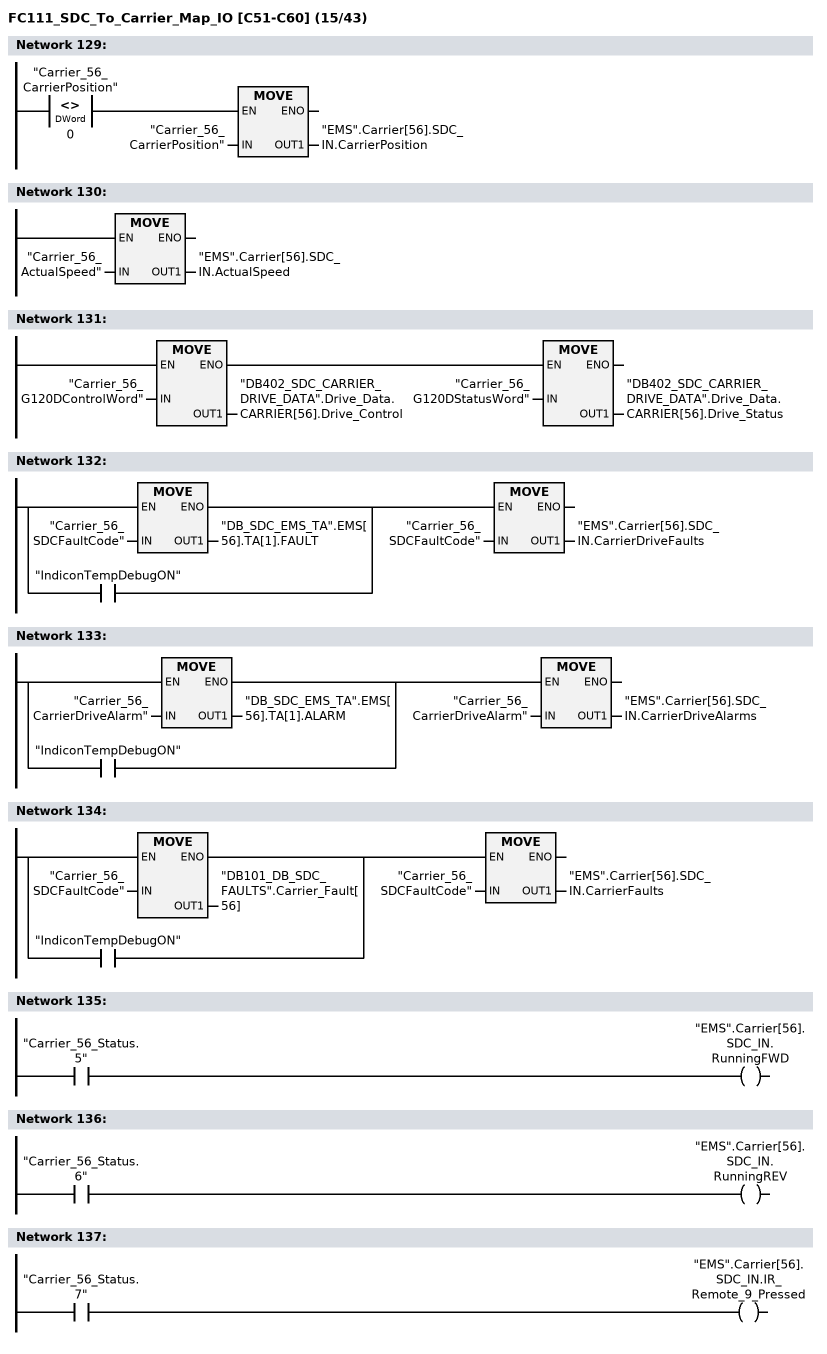
   RUNG wire#powerrail
      { S7_Templates := "SrcType := DWord" } NE_Contact(in1 := "Carrier_56_CarrierPosition", in2 := 0)
      Move(in := "Carrier_56_CarrierPosition", out1 => "EMS".Carrier[56].SDC_IN.CarrierPosition)
   END_RUNG
   // the same network as SCL:
   IF "Carrier_56_CarrierPosition" <> 0 THEN
       "EMS".Carrier[56].SDC_IN.CarrierPosition := "Carrier_56_CarrierPosition";
   END_IF;
END_REGION

REGION Network 130
   RUNG wire#powerrail
      Move(in := "Carrier_56_ActualSpeed", out1 => "EMS".Carrier[56].SDC_IN.ActualSpeed)
   END_RUNG
   // the same network as SCL:
   "EMS".Carrier[56].SDC_IN.ActualSpeed := "Carrier_56_ActualSpeed";
END_REGION

REGION Network 131
   RUNG wire#powerrail
      Move(in := "Carrier_56_G120DControlWord", out1 => "DB402_SDC_CARRIER_DRIVE_DATA".Drive_Data.CARRIER[56].Drive_Control)
      Move(in := "Carrier_56_G120DStatusWord", out1 => "DB402_SDC_CARRIER_DRIVE_DATA".Drive_Data.CARRIER[56].Drive_Status)
   END_RUNG
   // the same network as SCL:
   "DB402_SDC_CARRIER_DRIVE_DATA".Drive_Data.CARRIER[56].Drive_Control := "Carrier_56_G120DControlWord";
   "DB402_SDC_CARRIER_DRIVE_DATA".Drive_Data.CARRIER[56].Drive_Status := "Carrier_56_G120DStatusWord";
END_REGION

REGION Network 132
   RUNG wire#powerrail
      Move(in := "Carrier_56_SDCFaultCode", out1 => "DB_SDC_EMS_TA".EMS[56].TA[1].FAULT)
      wire#w1
      Move(in := "Carrier_56_SDCFaultCode", out1 => "EMS".Carrier[56].SDC_IN.CarrierDriveFaults)
   END_RUNG
   RUNG wire#powerrail
      Contact( "IndiconTempDebugON" )
   END_RUNG wire#w1
   // the same network as SCL:
   "DB_SDC_EMS_TA".EMS[56].TA[1].FAULT := "Carrier_56_SDCFaultCode";
   IF TRUE OR "IndiconTempDebugON" THEN
       "EMS".Carrier[56].SDC_IN.CarrierDriveFaults := "Carrier_56_SDCFaultCode";
   END_IF;
END_REGION

REGION Network 133
   RUNG wire#powerrail
      Move(in := "Carrier_56_CarrierDriveAlarm", out1 => "DB_SDC_EMS_TA".EMS[56].TA[1].ALARM)
      wire#w1
      Move(in := "Carrier_56_CarrierDriveAlarm", out1 => "EMS".Carrier[56].SDC_IN.CarrierDriveAlarms)
   END_RUNG
   RUNG wire#powerrail
      Contact( "IndiconTempDebugON" )
   END_RUNG wire#w1
   // the same network as SCL:
   "DB_SDC_EMS_TA".EMS[56].TA[1].ALARM := "Carrier_56_CarrierDriveAlarm";
   IF TRUE OR "IndiconTempDebugON" THEN
       "EMS".Carrier[56].SDC_IN.CarrierDriveAlarms := "Carrier_56_CarrierDriveAlarm";
   END_IF;
END_REGION

REGION Network 134
   RUNG wire#powerrail
      Move(in := "Carrier_56_SDCFaultCode", out1 => "DB101_DB_SDC_FAULTS".Carrier_Fault[56])
      wire#w1
      Move(in := "Carrier_56_SDCFaultCode", out1 => "EMS".Carrier[56].SDC_IN.CarrierFaults)
   END_RUNG
   RUNG wire#powerrail
      Contact( "IndiconTempDebugON" )
   END_RUNG wire#w1
   // the same network as SCL:
   "DB101_DB_SDC_FAULTS".Carrier_Fault[56] := "Carrier_56_SDCFaultCode";
   IF TRUE OR "IndiconTempDebugON" THEN
       "EMS".Carrier[56].SDC_IN.CarrierFaults := "Carrier_56_SDCFaultCode";
   END_IF;
END_REGION

REGION Network 135
   RUNG wire#powerrail
      Contact( "Carrier_56_Status.5" )
      Coil( "EMS".Carrier[56].SDC_IN.RunningFWD )
   END_RUNG
   // the same network as SCL:
   "EMS".Carrier[56].SDC_IN.RunningFWD := "Carrier_56_Status.5";
END_REGION

REGION Network 136
   RUNG wire#powerrail
      Contact( "Carrier_56_Status.6" )
      Coil( "EMS".Carrier[56].SDC_IN.RunningREV )
   END_RUNG
   // the same network as SCL:
   "EMS".Carrier[56].SDC_IN.RunningREV := "Carrier_56_Status.6";
END_REGION

REGION Network 137
   RUNG wire#powerrail
      Contact( "Carrier_56_Status.7" )
      Coil( "EMS".Carrier[56].SDC_IN.IR_Remote_9_Pressed )
   END_RUNG
   // the same network as SCL:
   "EMS".Carrier[56].SDC_IN.IR_Remote_9_Pressed := "Carrier_56_Status.7";
END_REGION

REGION Network 138
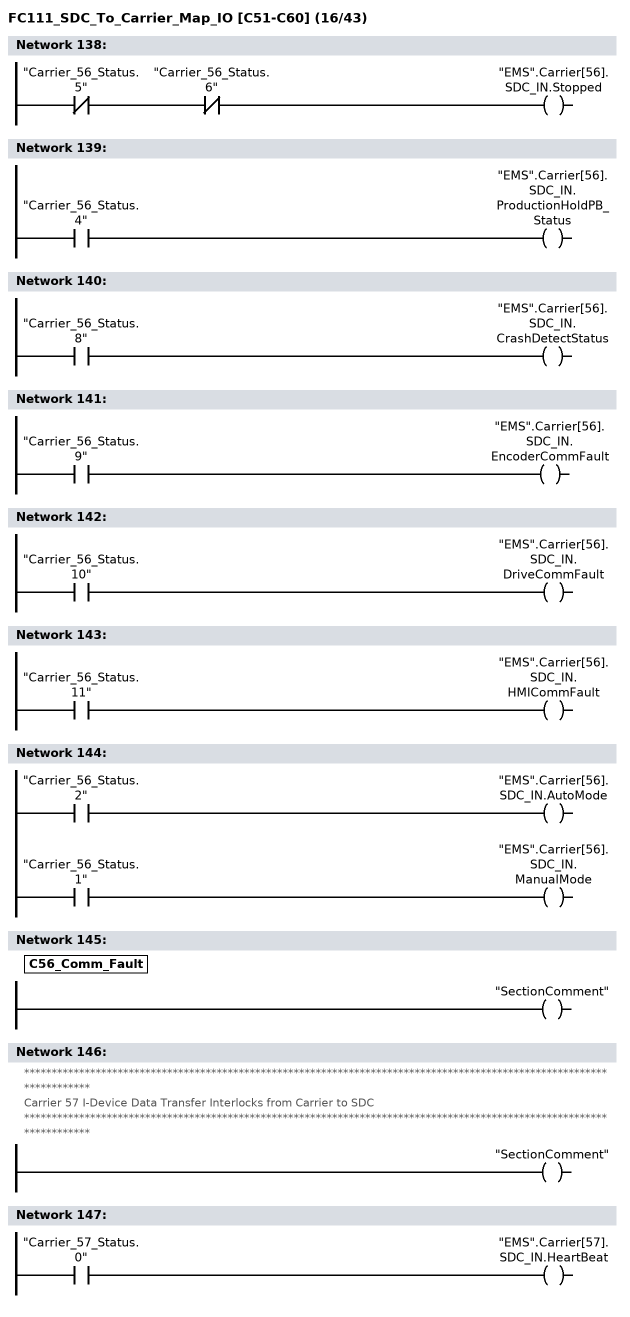
   RUNG wire#powerrail
      I_Contact( "Carrier_56_Status.5" )
      I_Contact( "Carrier_56_Status.6" )
      Coil( "EMS".Carrier[56].SDC_IN.Stopped )
   END_RUNG
   // the same network as SCL:
   "EMS".Carrier[56].SDC_IN.Stopped := NOT "Carrier_56_Status.5" AND NOT "Carrier_56_Status.6";
END_REGION

REGION Network 139
   RUNG wire#powerrail
      Contact( "Carrier_56_Status.4" )
      Coil( "EMS".Carrier[56].SDC_IN.ProductionHoldPB_Status )
   END_RUNG
   // the same network as SCL:
   "EMS".Carrier[56].SDC_IN.ProductionHoldPB_Status := "Carrier_56_Status.4";
END_REGION

REGION Network 140
   RUNG wire#powerrail
      Contact( "Carrier_56_Status.8" )
      Coil( "EMS".Carrier[56].SDC_IN.CrashDetectStatus )
   END_RUNG
   // the same network as SCL:
   "EMS".Carrier[56].SDC_IN.CrashDetectStatus := "Carrier_56_Status.8";
END_REGION

REGION Network 141
   RUNG wire#powerrail
      Contact( "Carrier_56_Status.9" )
      Coil( "EMS".Carrier[56].SDC_IN.EncoderCommFault )
   END_RUNG
   // the same network as SCL:
   "EMS".Carrier[56].SDC_IN.EncoderCommFault := "Carrier_56_Status.9";
END_REGION

REGION Network 142
   RUNG wire#powerrail
      Contact( "Carrier_56_Status.10" )
      Coil( "EMS".Carrier[56].SDC_IN.DriveCommFault )
   END_RUNG
   // the same network as SCL:
   "EMS".Carrier[56].SDC_IN.DriveCommFault := "Carrier_56_Status.10";
END_REGION

REGION Network 143
   RUNG wire#powerrail
      Contact( "Carrier_56_Status.11" )
      Coil( "EMS".Carrier[56].SDC_IN.HMICommFault )
   END_RUNG
   // the same network as SCL:
   "EMS".Carrier[56].SDC_IN.HMICommFault := "Carrier_56_Status.11";
END_REGION

REGION Network 144
   RUNG wire#powerrail
      Contact( "Carrier_56_Status.2" )
      Coil( "EMS".Carrier[56].SDC_IN.AutoMode )
   END_RUNG
   RUNG wire#powerrail
      Contact( "Carrier_56_Status.1" )
      Coil( "EMS".Carrier[56].SDC_IN.ManualMode )
   END_RUNG
   // the same network as SCL:
   "EMS".Carrier[56].SDC_IN.AutoMode := "Carrier_56_Status.2";
   "EMS".Carrier[56].SDC_IN.ManualMode := "Carrier_56_Status.1";
END_REGION

REGION Network 145
   Label( C56_Comm_Fault )
   RUNG wire#powerrail
      Coil( "SectionComment" )
   END_RUNG
   // the same network as SCL:
   C56_Comm_Fault:
   "SectionComment" := TRUE;
END_REGION

REGION Network 146
   // **********************************************************************************************************************
   // 
   // Carrier 57 I-Device Data Transfer Interlocks from Carrier to SDC
   // 
   // **********************************************************************************************************************
   RUNG wire#powerrail
      Coil( "SectionComment" )
   END_RUNG
   // the same network as SCL:
   "SectionComment" := TRUE;
END_REGION

REGION Network 147
   RUNG wire#powerrail
      Contact( "Carrier_57_Status.0" )
      Coil( "EMS".Carrier[57].SDC_IN.HeartBeat )
   END_RUNG
   // the same network as SCL:
   "EMS".Carrier[57].SDC_IN.HeartBeat := "Carrier_57_Status.0";
END_REGION

REGION Network 148
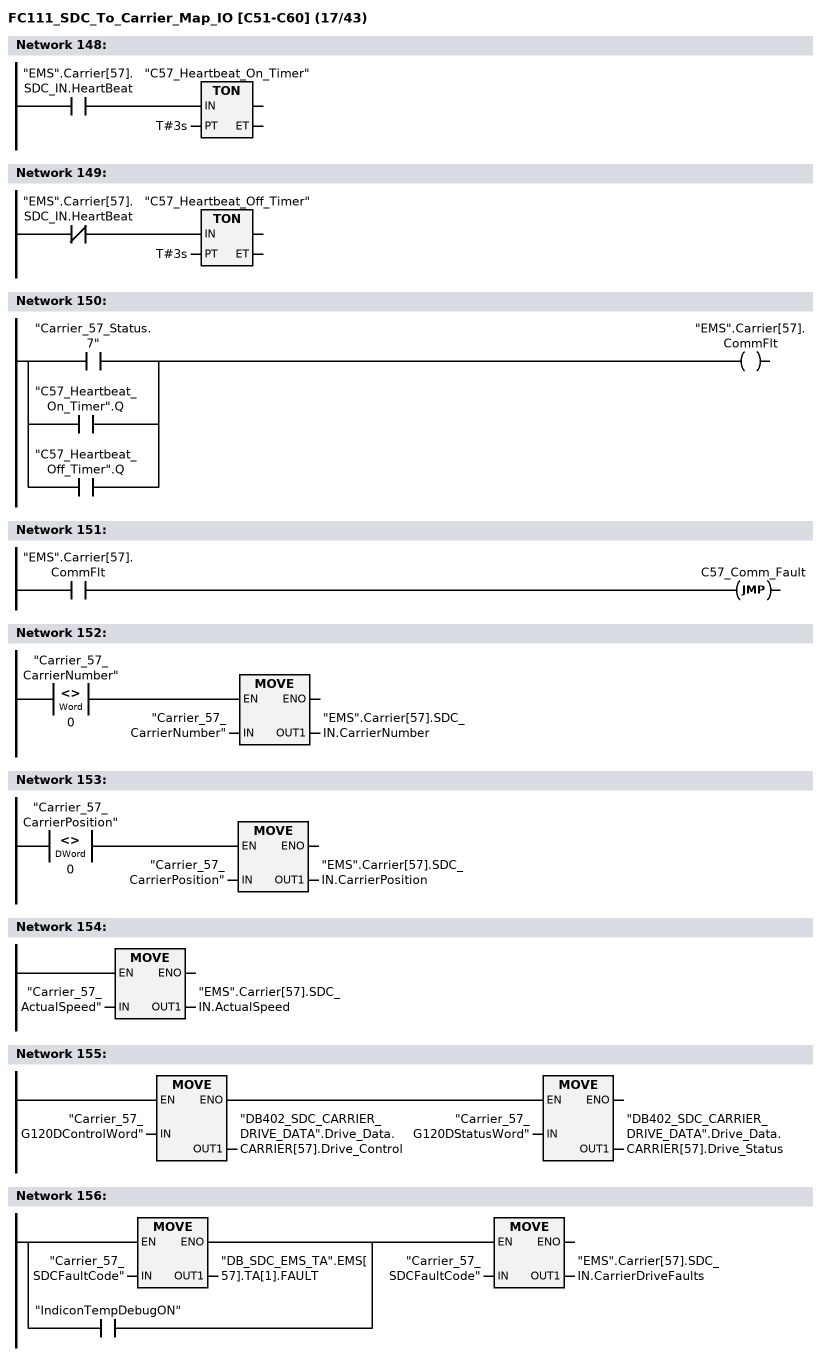
   "C57_Heartbeat_On_Timer".TON(IN := "EMS".Carrier[57].SDC_IN.HeartBeat, PT := T#3s);
END_REGION

REGION Network 149
   "C57_Heartbeat_Off_Timer".TON(IN := NOT "EMS".Carrier[57].SDC_IN.HeartBeat, PT := T#3s);
END_REGION

REGION Network 150
   RUNG wire#powerrail
      Contact( "Carrier_57_Status.7" )
      wire#w1
      Coil( "EMS".Carrier[57].CommFlt )
   END_RUNG
   RUNG wire#powerrail
      Contact( "C57_Heartbeat_On_Timer".Q )
   END_RUNG wire#w1
   RUNG wire#powerrail
      Contact( "C57_Heartbeat_Off_Timer".Q )
   END_RUNG wire#w1
   // the same network as SCL:
   "EMS".Carrier[57].CommFlt := "Carrier_57_Status.7" OR "C57_Heartbeat_On_Timer".Q OR "C57_Heartbeat_Off_Timer".Q;
END_REGION

REGION Network 151
   RUNG wire#powerrail
      Contact( "EMS".Carrier[57].CommFlt )
      JumpCoil( C57_Comm_Fault )
   END_RUNG
   // the same network as SCL:
   IF "EMS".Carrier[57].CommFlt THEN GOTO C57_Comm_Fault; END_IF;
END_REGION

REGION Network 152
   RUNG wire#powerrail
      { S7_Templates := "SrcType := Word" } NE_Contact(in1 := "Carrier_57_CarrierNumber", in2 := 0)
      Move(in := "Carrier_57_CarrierNumber", out1 => "EMS".Carrier[57].SDC_IN.CarrierNumber)
   END_RUNG
   // the same network as SCL:
   IF "Carrier_57_CarrierNumber" <> 0 THEN
       "EMS".Carrier[57].SDC_IN.CarrierNumber := "Carrier_57_CarrierNumber";
   END_IF;
END_REGION

REGION Network 153
   RUNG wire#powerrail
      { S7_Templates := "SrcType := DWord" } NE_Contact(in1 := "Carrier_57_CarrierPosition", in2 := 0)
      Move(in := "Carrier_57_CarrierPosition", out1 => "EMS".Carrier[57].SDC_IN.CarrierPosition)
   END_RUNG
   // the same network as SCL:
   IF "Carrier_57_CarrierPosition" <> 0 THEN
       "EMS".Carrier[57].SDC_IN.CarrierPosition := "Carrier_57_CarrierPosition";
   END_IF;
END_REGION

REGION Network 154
   RUNG wire#powerrail
      Move(in := "Carrier_57_ActualSpeed", out1 => "EMS".Carrier[57].SDC_IN.ActualSpeed)
   END_RUNG
   // the same network as SCL:
   "EMS".Carrier[57].SDC_IN.ActualSpeed := "Carrier_57_ActualSpeed";
END_REGION

REGION Network 155
   RUNG wire#powerrail
      Move(in := "Carrier_57_G120DControlWord", out1 => "DB402_SDC_CARRIER_DRIVE_DATA".Drive_Data.CARRIER[57].Drive_Control)
      Move(in := "Carrier_57_G120DStatusWord", out1 => "DB402_SDC_CARRIER_DRIVE_DATA".Drive_Data.CARRIER[57].Drive_Status)
   END_RUNG
   // the same network as SCL:
   "DB402_SDC_CARRIER_DRIVE_DATA".Drive_Data.CARRIER[57].Drive_Control := "Carrier_57_G120DControlWord";
   "DB402_SDC_CARRIER_DRIVE_DATA".Drive_Data.CARRIER[57].Drive_Status := "Carrier_57_G120DStatusWord";
END_REGION

REGION Network 156
   RUNG wire#powerrail
      Move(in := "Carrier_57_SDCFaultCode", out1 => "DB_SDC_EMS_TA".EMS[57].TA[1].FAULT)
      wire#w1
      Move(in := "Carrier_57_SDCFaultCode", out1 => "EMS".Carrier[57].SDC_IN.CarrierDriveFaults)
   END_RUNG
   RUNG wire#powerrail
      Contact( "IndiconTempDebugON" )
   END_RUNG wire#w1
   // the same network as SCL:
   "DB_SDC_EMS_TA".EMS[57].TA[1].FAULT := "Carrier_57_SDCFaultCode";
   IF TRUE OR "IndiconTempDebugON" THEN
       "EMS".Carrier[57].SDC_IN.CarrierDriveFaults := "Carrier_57_SDCFaultCode";
   END_IF;
END_REGION

REGION Network 157
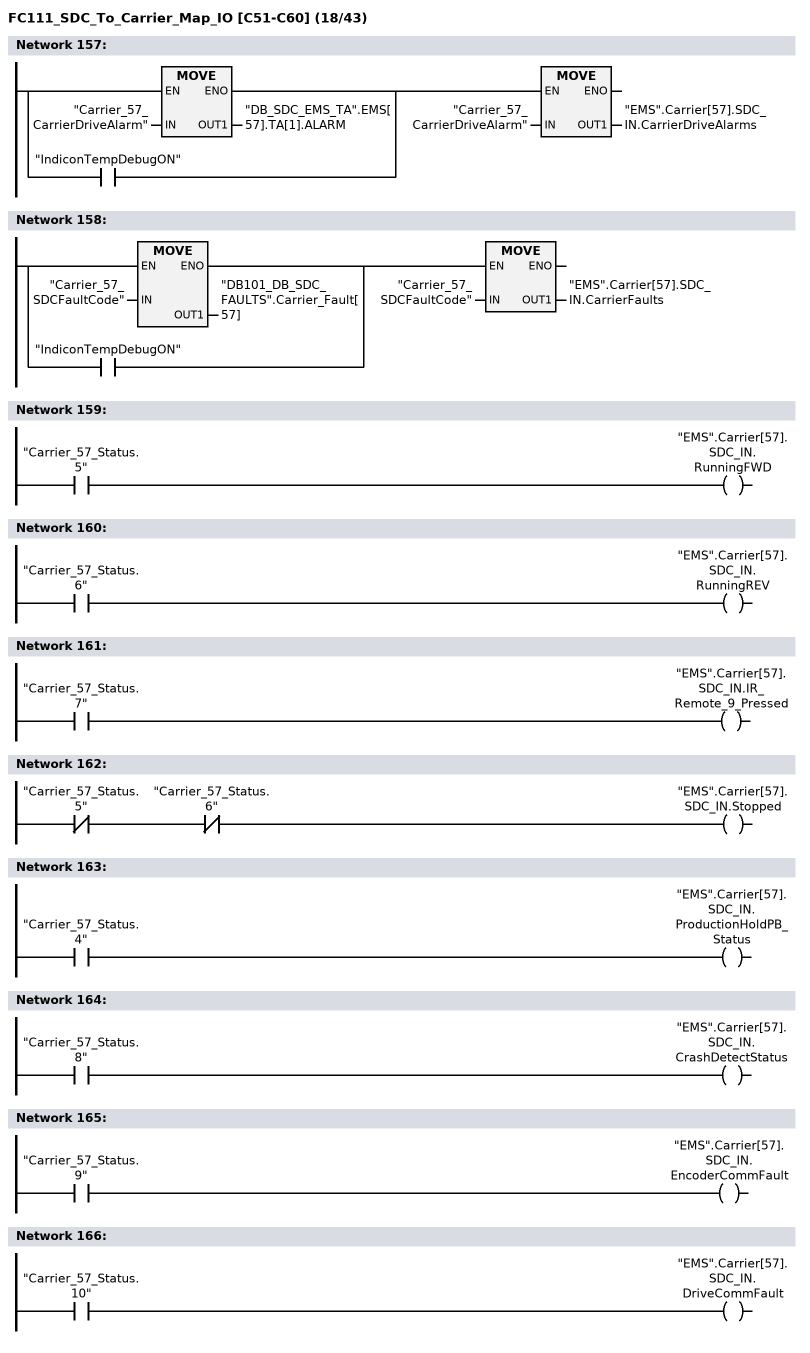
   RUNG wire#powerrail
      Move(in := "Carrier_57_CarrierDriveAlarm", out1 => "DB_SDC_EMS_TA".EMS[57].TA[1].ALARM)
      wire#w1
      Move(in := "Carrier_57_CarrierDriveAlarm", out1 => "EMS".Carrier[57].SDC_IN.CarrierDriveAlarms)
   END_RUNG
   RUNG wire#powerrail
      Contact( "IndiconTempDebugON" )
   END_RUNG wire#w1
   // the same network as SCL:
   "DB_SDC_EMS_TA".EMS[57].TA[1].ALARM := "Carrier_57_CarrierDriveAlarm";
   IF TRUE OR "IndiconTempDebugON" THEN
       "EMS".Carrier[57].SDC_IN.CarrierDriveAlarms := "Carrier_57_CarrierDriveAlarm";
   END_IF;
END_REGION

REGION Network 158
   RUNG wire#powerrail
      Move(in := "Carrier_57_SDCFaultCode", out1 => "DB101_DB_SDC_FAULTS".Carrier_Fault[57])
      wire#w1
      Move(in := "Carrier_57_SDCFaultCode", out1 => "EMS".Carrier[57].SDC_IN.CarrierFaults)
   END_RUNG
   RUNG wire#powerrail
      Contact( "IndiconTempDebugON" )
   END_RUNG wire#w1
   // the same network as SCL:
   "DB101_DB_SDC_FAULTS".Carrier_Fault[57] := "Carrier_57_SDCFaultCode";
   IF TRUE OR "IndiconTempDebugON" THEN
       "EMS".Carrier[57].SDC_IN.CarrierFaults := "Carrier_57_SDCFaultCode";
   END_IF;
END_REGION

REGION Network 159
   RUNG wire#powerrail
      Contact( "Carrier_57_Status.5" )
      Coil( "EMS".Carrier[57].SDC_IN.RunningFWD )
   END_RUNG
   // the same network as SCL:
   "EMS".Carrier[57].SDC_IN.RunningFWD := "Carrier_57_Status.5";
END_REGION

REGION Network 160
   RUNG wire#powerrail
      Contact( "Carrier_57_Status.6" )
      Coil( "EMS".Carrier[57].SDC_IN.RunningREV )
   END_RUNG
   // the same network as SCL:
   "EMS".Carrier[57].SDC_IN.RunningREV := "Carrier_57_Status.6";
END_REGION

REGION Network 161
   RUNG wire#powerrail
      Contact( "Carrier_57_Status.7" )
      Coil( "EMS".Carrier[57].SDC_IN.IR_Remote_9_Pressed )
   END_RUNG
   // the same network as SCL:
   "EMS".Carrier[57].SDC_IN.IR_Remote_9_Pressed := "Carrier_57_Status.7";
END_REGION

REGION Network 162
   RUNG wire#powerrail
      I_Contact( "Carrier_57_Status.5" )
      I_Contact( "Carrier_57_Status.6" )
      Coil( "EMS".Carrier[57].SDC_IN.Stopped )
   END_RUNG
   // the same network as SCL:
   "EMS".Carrier[57].SDC_IN.Stopped := NOT "Carrier_57_Status.5" AND NOT "Carrier_57_Status.6";
END_REGION

REGION Network 163
   RUNG wire#powerrail
      Contact( "Carrier_57_Status.4" )
      Coil( "EMS".Carrier[57].SDC_IN.ProductionHoldPB_Status )
   END_RUNG
   // the same network as SCL:
   "EMS".Carrier[57].SDC_IN.ProductionHoldPB_Status := "Carrier_57_Status.4";
END_REGION

REGION Network 164
   RUNG wire#powerrail
      Contact( "Carrier_57_Status.8" )
      Coil( "EMS".Carrier[57].SDC_IN.CrashDetectStatus )
   END_RUNG
   // the same network as SCL:
   "EMS".Carrier[57].SDC_IN.CrashDetectStatus := "Carrier_57_Status.8";
END_REGION

REGION Network 165
   RUNG wire#powerrail
      Contact( "Carrier_57_Status.9" )
      Coil( "EMS".Carrier[57].SDC_IN.EncoderCommFault )
   END_RUNG
   // the same network as SCL:
   "EMS".Carrier[57].SDC_IN.EncoderCommFault := "Carrier_57_Status.9";
END_REGION

REGION Network 166
   RUNG wire#powerrail
      Contact( "Carrier_57_Status.10" )
      Coil( "EMS".Carrier[57].SDC_IN.DriveCommFault )
   END_RUNG
   // the same network as SCL:
   "EMS".Carrier[57].SDC_IN.DriveCommFault := "Carrier_57_Status.10";
END_REGION

REGION Network 167
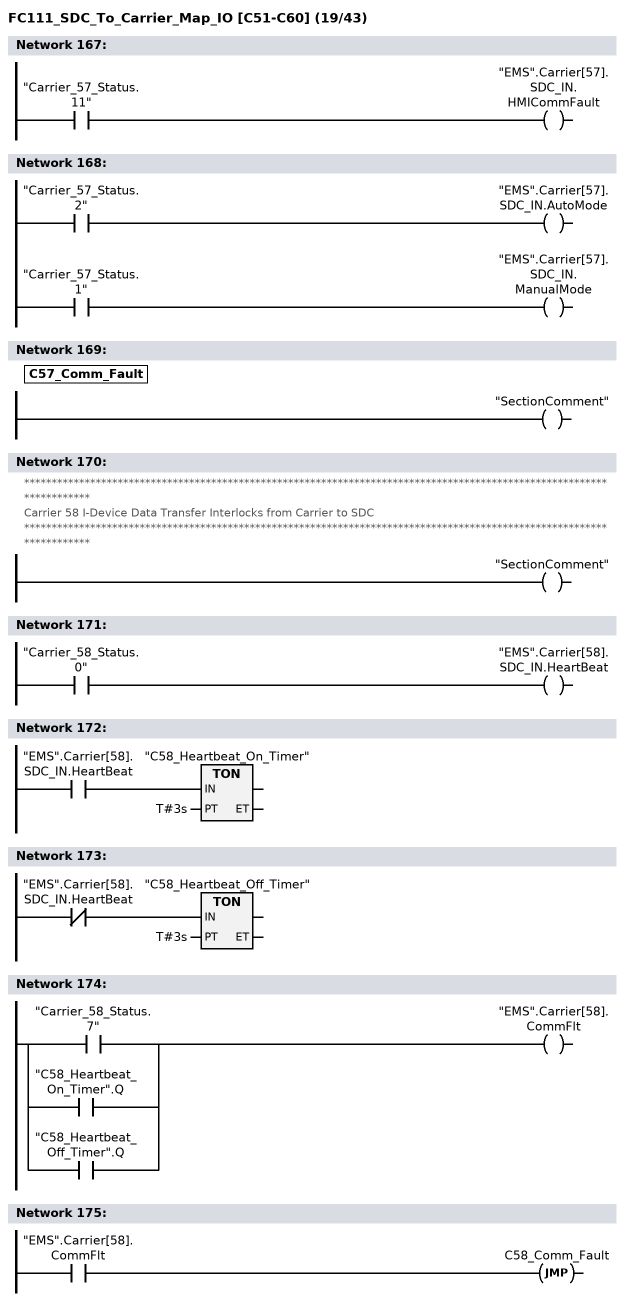
   RUNG wire#powerrail
      Contact( "Carrier_57_Status.11" )
      Coil( "EMS".Carrier[57].SDC_IN.HMICommFault )
   END_RUNG
   // the same network as SCL:
   "EMS".Carrier[57].SDC_IN.HMICommFault := "Carrier_57_Status.11";
END_REGION

REGION Network 168
   RUNG wire#powerrail
      Contact( "Carrier_57_Status.2" )
      Coil( "EMS".Carrier[57].SDC_IN.AutoMode )
   END_RUNG
   RUNG wire#powerrail
      Contact( "Carrier_57_Status.1" )
      Coil( "EMS".Carrier[57].SDC_IN.ManualMode )
   END_RUNG
   // the same network as SCL:
   "EMS".Carrier[57].SDC_IN.AutoMode := "Carrier_57_Status.2";
   "EMS".Carrier[57].SDC_IN.ManualMode := "Carrier_57_Status.1";
END_REGION

REGION Network 169
   Label( C57_Comm_Fault )
   RUNG wire#powerrail
      Coil( "SectionComment" )
   END_RUNG
   // the same network as SCL:
   C57_Comm_Fault:
   "SectionComment" := TRUE;
END_REGION

REGION Network 170
   // **********************************************************************************************************************
   // 
   // Carrier 58 I-Device Data Transfer Interlocks from Carrier to SDC
   // 
   // **********************************************************************************************************************
   RUNG wire#powerrail
      Coil( "SectionComment" )
   END_RUNG
   // the same network as SCL:
   "SectionComment" := TRUE;
END_REGION

REGION Network 171
   RUNG wire#powerrail
      Contact( "Carrier_58_Status.0" )
      Coil( "EMS".Carrier[58].SDC_IN.HeartBeat )
   END_RUNG
   // the same network as SCL:
   "EMS".Carrier[58].SDC_IN.HeartBeat := "Carrier_58_Status.0";
END_REGION

REGION Network 172
   "C58_Heartbeat_On_Timer".TON(IN := "EMS".Carrier[58].SDC_IN.HeartBeat, PT := T#3s);
END_REGION

REGION Network 173
   "C58_Heartbeat_Off_Timer".TON(IN := NOT "EMS".Carrier[58].SDC_IN.HeartBeat, PT := T#3s);
END_REGION

REGION Network 174
   RUNG wire#powerrail
      Contact( "Carrier_58_Status.7" )
      wire#w1
      Coil( "EMS".Carrier[58].CommFlt )
   END_RUNG
   RUNG wire#powerrail
      Contact( "C58_Heartbeat_On_Timer".Q )
   END_RUNG wire#w1
   RUNG wire#powerrail
      Contact( "C58_Heartbeat_Off_Timer".Q )
   END_RUNG wire#w1
   // the same network as SCL:
   "EMS".Carrier[58].CommFlt := "Carrier_58_Status.7" OR "C58_Heartbeat_On_Timer".Q OR "C58_Heartbeat_Off_Timer".Q;
END_REGION

REGION Network 175
   RUNG wire#powerrail
      Contact( "EMS".Carrier[58].CommFlt )
      JumpCoil( C58_Comm_Fault )
   END_RUNG
   // the same network as SCL:
   IF "EMS".Carrier[58].CommFlt THEN GOTO C58_Comm_Fault; END_IF;
END_REGION

REGION Network 176
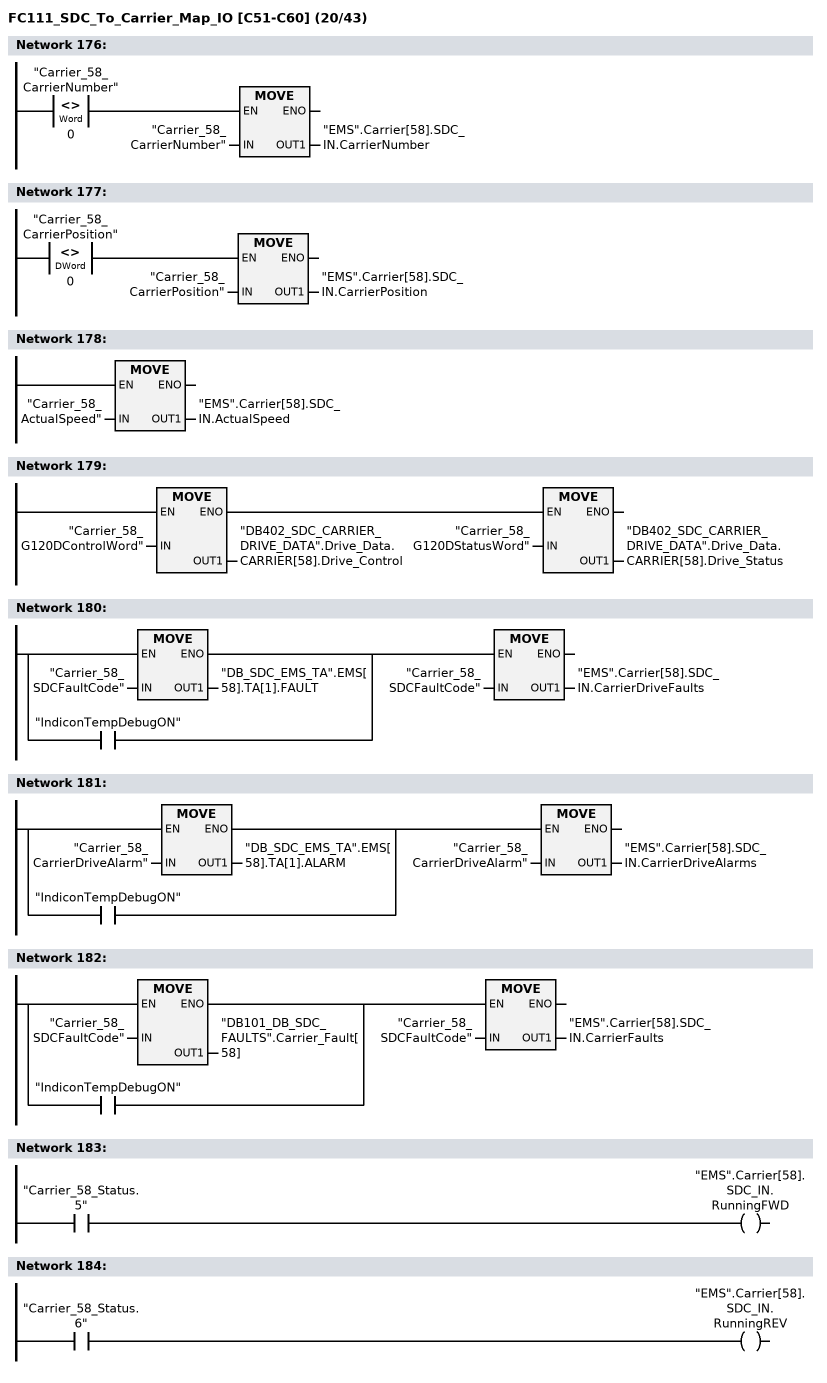
   RUNG wire#powerrail
      { S7_Templates := "SrcType := Word" } NE_Contact(in1 := "Carrier_58_CarrierNumber", in2 := 0)
      Move(in := "Carrier_58_CarrierNumber", out1 => "EMS".Carrier[58].SDC_IN.CarrierNumber)
   END_RUNG
   // the same network as SCL:
   IF "Carrier_58_CarrierNumber" <> 0 THEN
       "EMS".Carrier[58].SDC_IN.CarrierNumber := "Carrier_58_CarrierNumber";
   END_IF;
END_REGION

REGION Network 177
   RUNG wire#powerrail
      { S7_Templates := "SrcType := DWord" } NE_Contact(in1 := "Carrier_58_CarrierPosition", in2 := 0)
      Move(in := "Carrier_58_CarrierPosition", out1 => "EMS".Carrier[58].SDC_IN.CarrierPosition)
   END_RUNG
   // the same network as SCL:
   IF "Carrier_58_CarrierPosition" <> 0 THEN
       "EMS".Carrier[58].SDC_IN.CarrierPosition := "Carrier_58_CarrierPosition";
   END_IF;
END_REGION

REGION Network 178
   RUNG wire#powerrail
      Move(in := "Carrier_58_ActualSpeed", out1 => "EMS".Carrier[58].SDC_IN.ActualSpeed)
   END_RUNG
   // the same network as SCL:
   "EMS".Carrier[58].SDC_IN.ActualSpeed := "Carrier_58_ActualSpeed";
END_REGION

REGION Network 179
   RUNG wire#powerrail
      Move(in := "Carrier_58_G120DControlWord", out1 => "DB402_SDC_CARRIER_DRIVE_DATA".Drive_Data.CARRIER[58].Drive_Control)
      Move(in := "Carrier_58_G120DStatusWord", out1 => "DB402_SDC_CARRIER_DRIVE_DATA".Drive_Data.CARRIER[58].Drive_Status)
   END_RUNG
   // the same network as SCL:
   "DB402_SDC_CARRIER_DRIVE_DATA".Drive_Data.CARRIER[58].Drive_Control := "Carrier_58_G120DControlWord";
   "DB402_SDC_CARRIER_DRIVE_DATA".Drive_Data.CARRIER[58].Drive_Status := "Carrier_58_G120DStatusWord";
END_REGION

REGION Network 180
   RUNG wire#powerrail
      Move(in := "Carrier_58_SDCFaultCode", out1 => "DB_SDC_EMS_TA".EMS[58].TA[1].FAULT)
      wire#w1
      Move(in := "Carrier_58_SDCFaultCode", out1 => "EMS".Carrier[58].SDC_IN.CarrierDriveFaults)
   END_RUNG
   RUNG wire#powerrail
      Contact( "IndiconTempDebugON" )
   END_RUNG wire#w1
   // the same network as SCL:
   "DB_SDC_EMS_TA".EMS[58].TA[1].FAULT := "Carrier_58_SDCFaultCode";
   IF TRUE OR "IndiconTempDebugON" THEN
       "EMS".Carrier[58].SDC_IN.CarrierDriveFaults := "Carrier_58_SDCFaultCode";
   END_IF;
END_REGION

REGION Network 181
   RUNG wire#powerrail
      Move(in := "Carrier_58_CarrierDriveAlarm", out1 => "DB_SDC_EMS_TA".EMS[58].TA[1].ALARM)
      wire#w1
      Move(in := "Carrier_58_CarrierDriveAlarm", out1 => "EMS".Carrier[58].SDC_IN.CarrierDriveAlarms)
   END_RUNG
   RUNG wire#powerrail
      Contact( "IndiconTempDebugON" )
   END_RUNG wire#w1
   // the same network as SCL:
   "DB_SDC_EMS_TA".EMS[58].TA[1].ALARM := "Carrier_58_CarrierDriveAlarm";
   IF TRUE OR "IndiconTempDebugON" THEN
       "EMS".Carrier[58].SDC_IN.CarrierDriveAlarms := "Carrier_58_CarrierDriveAlarm";
   END_IF;
END_REGION

REGION Network 182
   RUNG wire#powerrail
      Move(in := "Carrier_58_SDCFaultCode", out1 => "DB101_DB_SDC_FAULTS".Carrier_Fault[58])
      wire#w1
      Move(in := "Carrier_58_SDCFaultCode", out1 => "EMS".Carrier[58].SDC_IN.CarrierFaults)
   END_RUNG
   RUNG wire#powerrail
      Contact( "IndiconTempDebugON" )
   END_RUNG wire#w1
   // the same network as SCL:
   "DB101_DB_SDC_FAULTS".Carrier_Fault[58] := "Carrier_58_SDCFaultCode";
   IF TRUE OR "IndiconTempDebugON" THEN
       "EMS".Carrier[58].SDC_IN.CarrierFaults := "Carrier_58_SDCFaultCode";
   END_IF;
END_REGION

REGION Network 183
   RUNG wire#powerrail
      Contact( "Carrier_58_Status.5" )
      Coil( "EMS".Carrier[58].SDC_IN.RunningFWD )
   END_RUNG
   // the same network as SCL:
   "EMS".Carrier[58].SDC_IN.RunningFWD := "Carrier_58_Status.5";
END_REGION

REGION Network 184
   RUNG wire#powerrail
      Contact( "Carrier_58_Status.6" )
      Coil( "EMS".Carrier[58].SDC_IN.RunningREV )
   END_RUNG
   // the same network as SCL:
   "EMS".Carrier[58].SDC_IN.RunningREV := "Carrier_58_Status.6";
END_REGION

REGION Network 185
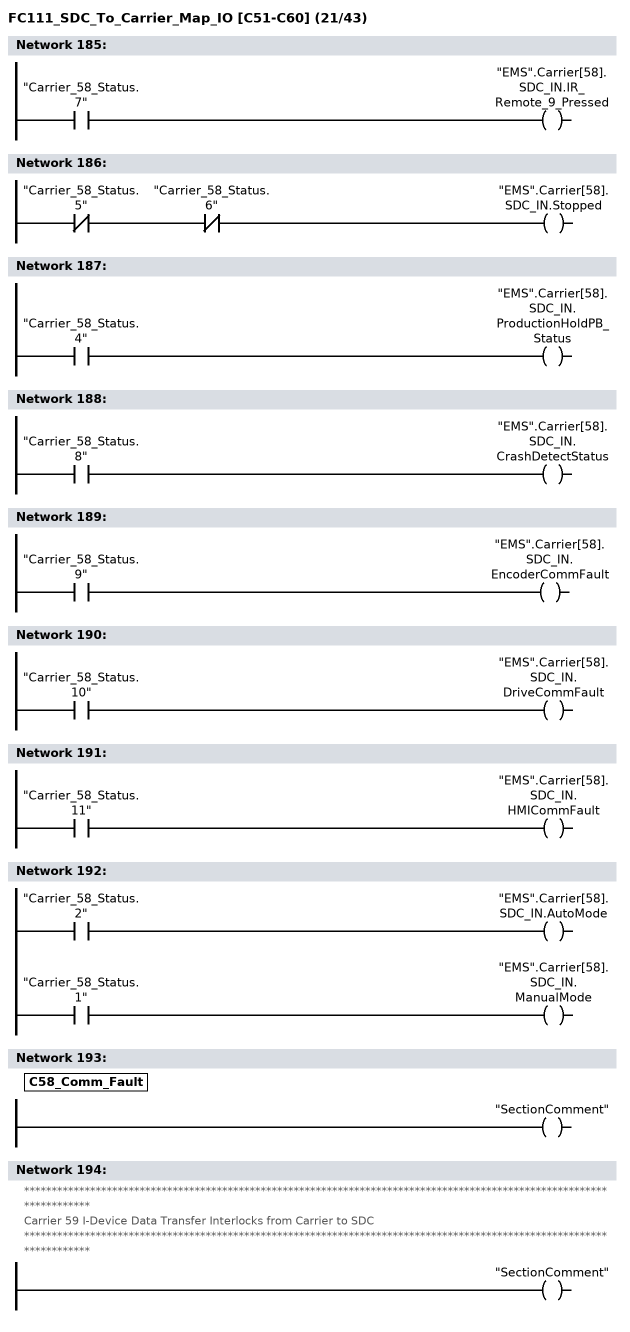
   RUNG wire#powerrail
      Contact( "Carrier_58_Status.7" )
      Coil( "EMS".Carrier[58].SDC_IN.IR_Remote_9_Pressed )
   END_RUNG
   // the same network as SCL:
   "EMS".Carrier[58].SDC_IN.IR_Remote_9_Pressed := "Carrier_58_Status.7";
END_REGION

REGION Network 186
   RUNG wire#powerrail
      I_Contact( "Carrier_58_Status.5" )
      I_Contact( "Carrier_58_Status.6" )
      Coil( "EMS".Carrier[58].SDC_IN.Stopped )
   END_RUNG
   // the same network as SCL:
   "EMS".Carrier[58].SDC_IN.Stopped := NOT "Carrier_58_Status.5" AND NOT "Carrier_58_Status.6";
END_REGION

REGION Network 187
   RUNG wire#powerrail
      Contact( "Carrier_58_Status.4" )
      Coil( "EMS".Carrier[58].SDC_IN.ProductionHoldPB_Status )
   END_RUNG
   // the same network as SCL:
   "EMS".Carrier[58].SDC_IN.ProductionHoldPB_Status := "Carrier_58_Status.4";
END_REGION

REGION Network 188
   RUNG wire#powerrail
      Contact( "Carrier_58_Status.8" )
      Coil( "EMS".Carrier[58].SDC_IN.CrashDetectStatus )
   END_RUNG
   // the same network as SCL:
   "EMS".Carrier[58].SDC_IN.CrashDetectStatus := "Carrier_58_Status.8";
END_REGION

REGION Network 189
   RUNG wire#powerrail
      Contact( "Carrier_58_Status.9" )
      Coil( "EMS".Carrier[58].SDC_IN.EncoderCommFault )
   END_RUNG
   // the same network as SCL:
   "EMS".Carrier[58].SDC_IN.EncoderCommFault := "Carrier_58_Status.9";
END_REGION

REGION Network 190
   RUNG wire#powerrail
      Contact( "Carrier_58_Status.10" )
      Coil( "EMS".Carrier[58].SDC_IN.DriveCommFault )
   END_RUNG
   // the same network as SCL:
   "EMS".Carrier[58].SDC_IN.DriveCommFault := "Carrier_58_Status.10";
END_REGION

REGION Network 191
   RUNG wire#powerrail
      Contact( "Carrier_58_Status.11" )
      Coil( "EMS".Carrier[58].SDC_IN.HMICommFault )
   END_RUNG
   // the same network as SCL:
   "EMS".Carrier[58].SDC_IN.HMICommFault := "Carrier_58_Status.11";
END_REGION

REGION Network 192
   RUNG wire#powerrail
      Contact( "Carrier_58_Status.2" )
      Coil( "EMS".Carrier[58].SDC_IN.AutoMode )
   END_RUNG
   RUNG wire#powerrail
      Contact( "Carrier_58_Status.1" )
      Coil( "EMS".Carrier[58].SDC_IN.ManualMode )
   END_RUNG
   // the same network as SCL:
   "EMS".Carrier[58].SDC_IN.AutoMode := "Carrier_58_Status.2";
   "EMS".Carrier[58].SDC_IN.ManualMode := "Carrier_58_Status.1";
END_REGION

REGION Network 193
   Label( C58_Comm_Fault )
   RUNG wire#powerrail
      Coil( "SectionComment" )
   END_RUNG
   // the same network as SCL:
   C58_Comm_Fault:
   "SectionComment" := TRUE;
END_REGION

REGION Network 194
   // **********************************************************************************************************************
   // 
   // Carrier 59 I-Device Data Transfer Interlocks from Carrier to SDC
   // 
   // **********************************************************************************************************************
   RUNG wire#powerrail
      Coil( "SectionComment" )
   END_RUNG
   // the same network as SCL:
   "SectionComment" := TRUE;
END_REGION

REGION Network 195
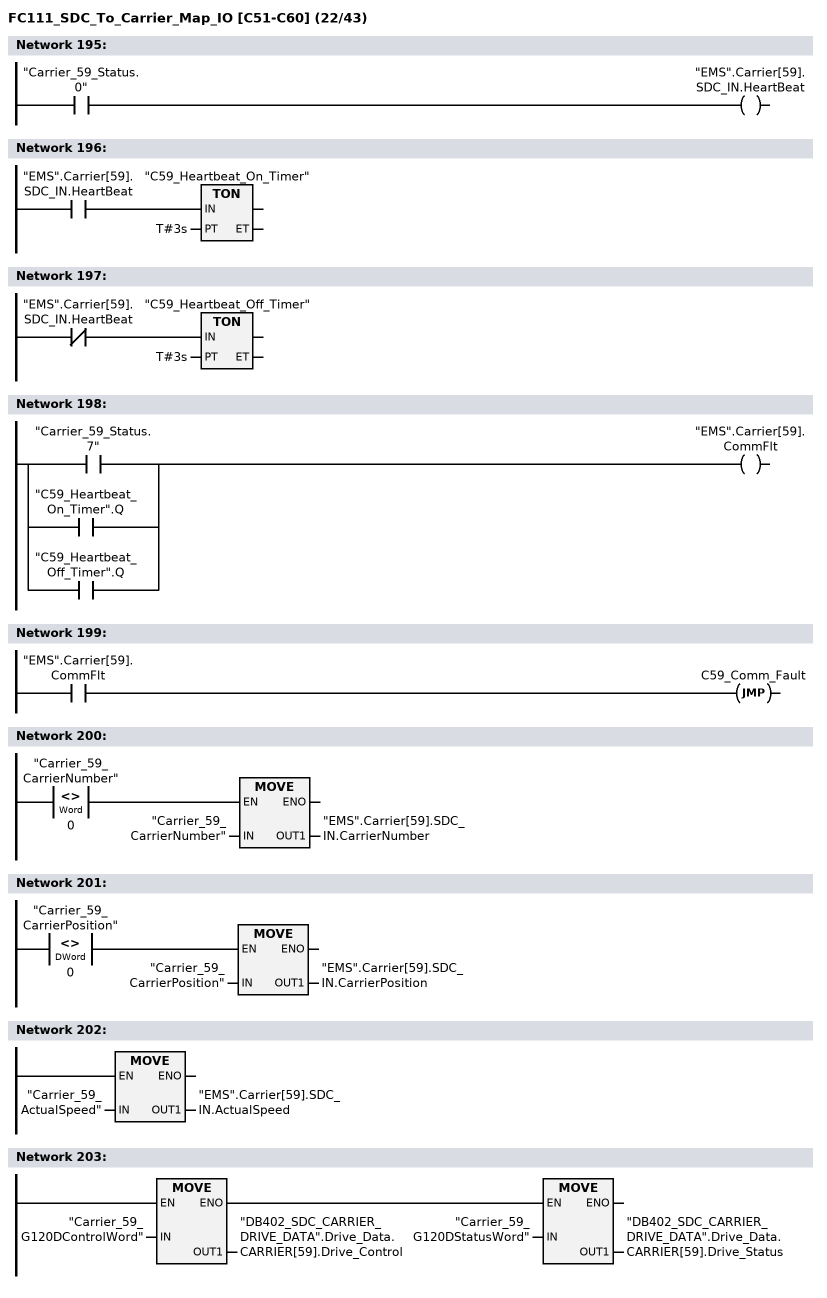
   RUNG wire#powerrail
      Contact( "Carrier_59_Status.0" )
      Coil( "EMS".Carrier[59].SDC_IN.HeartBeat )
   END_RUNG
   // the same network as SCL:
   "EMS".Carrier[59].SDC_IN.HeartBeat := "Carrier_59_Status.0";
END_REGION

REGION Network 196
   "C59_Heartbeat_On_Timer".TON(IN := "EMS".Carrier[59].SDC_IN.HeartBeat, PT := T#3s);
END_REGION

REGION Network 197
   "C59_Heartbeat_Off_Timer".TON(IN := NOT "EMS".Carrier[59].SDC_IN.HeartBeat, PT := T#3s);
END_REGION

REGION Network 198
   RUNG wire#powerrail
      Contact( "Carrier_59_Status.7" )
      wire#w1
      Coil( "EMS".Carrier[59].CommFlt )
   END_RUNG
   RUNG wire#powerrail
      Contact( "C59_Heartbeat_On_Timer".Q )
   END_RUNG wire#w1
   RUNG wire#powerrail
      Contact( "C59_Heartbeat_Off_Timer".Q )
   END_RUNG wire#w1
   // the same network as SCL:
   "EMS".Carrier[59].CommFlt := "Carrier_59_Status.7" OR "C59_Heartbeat_On_Timer".Q OR "C59_Heartbeat_Off_Timer".Q;
END_REGION

REGION Network 199
   RUNG wire#powerrail
      Contact( "EMS".Carrier[59].CommFlt )
      JumpCoil( C59_Comm_Fault )
   END_RUNG
   // the same network as SCL:
   IF "EMS".Carrier[59].CommFlt THEN GOTO C59_Comm_Fault; END_IF;
END_REGION

REGION Network 200
   RUNG wire#powerrail
      { S7_Templates := "SrcType := Word" } NE_Contact(in1 := "Carrier_59_CarrierNumber", in2 := 0)
      Move(in := "Carrier_59_CarrierNumber", out1 => "EMS".Carrier[59].SDC_IN.CarrierNumber)
   END_RUNG
   // the same network as SCL:
   IF "Carrier_59_CarrierNumber" <> 0 THEN
       "EMS".Carrier[59].SDC_IN.CarrierNumber := "Carrier_59_CarrierNumber";
   END_IF;
END_REGION

REGION Network 201
   RUNG wire#powerrail
      { S7_Templates := "SrcType := DWord" } NE_Contact(in1 := "Carrier_59_CarrierPosition", in2 := 0)
      Move(in := "Carrier_59_CarrierPosition", out1 => "EMS".Carrier[59].SDC_IN.CarrierPosition)
   END_RUNG
   // the same network as SCL:
   IF "Carrier_59_CarrierPosition" <> 0 THEN
       "EMS".Carrier[59].SDC_IN.CarrierPosition := "Carrier_59_CarrierPosition";
   END_IF;
END_REGION

REGION Network 202
   RUNG wire#powerrail
      Move(in := "Carrier_59_ActualSpeed", out1 => "EMS".Carrier[59].SDC_IN.ActualSpeed)
   END_RUNG
   // the same network as SCL:
   "EMS".Carrier[59].SDC_IN.ActualSpeed := "Carrier_59_ActualSpeed";
END_REGION

REGION Network 203
   RUNG wire#powerrail
      Move(in := "Carrier_59_G120DControlWord", out1 => "DB402_SDC_CARRIER_DRIVE_DATA".Drive_Data.CARRIER[59].Drive_Control)
      Move(in := "Carrier_59_G120DStatusWord", out1 => "DB402_SDC_CARRIER_DRIVE_DATA".Drive_Data.CARRIER[59].Drive_Status)
   END_RUNG
   // the same network as SCL:
   "DB402_SDC_CARRIER_DRIVE_DATA".Drive_Data.CARRIER[59].Drive_Control := "Carrier_59_G120DControlWord";
   "DB402_SDC_CARRIER_DRIVE_DATA".Drive_Data.CARRIER[59].Drive_Status := "Carrier_59_G120DStatusWord";
END_REGION

REGION Network 204
